FUNCTION_BLOCK "FB_BPSEthLink_V1.00"   // FB15, SCL
{ S7_Optimized_Access := 'TRUE' }
VERSION : 0.1
   VAR_INPUT
      IN_xBPSServerA : Bool;   // This istance is for BPS Server A
      IN_xCycleON : Bool;   // Cycle ON
      IN_xCycleONDel : Bool;   // Delayed cycle ON signal
      IN_xGeneralReset : Bool;   // General reset
      IN_xResetAlarms : Bool;   // Reset alarms
      IN_xFaultsEnabled : Bool;   // Faults enabled
      IN_xThisPLCActive : Bool;   // This PLC active
      IN_dLineSpeed_mm_min : DInt;   // Z301 speed [mm/min]
      IN_tStatusGeneral : Struct   // Status of general data
         dOptimizerMode : DInt;   // Optimizer mode (1=PLC 2=PC 3=Cullet)
         dExtOptSelected : DInt;   // External optimizer selected (1=PC A 2=PC B)
         dRibbonModality : DInt;   // Ribbon modality (1=Auto 4=Man)
         dAutoRibSelection : DInt;   // Automatic ribbon selection (0=Manual 1=Scanner 2=Camera)
         dTypeWanderSel : DInt;   // Wander type selection (1=Gross 2=Net)
         dActivePLC : DInt;   // Active PLC (1=PLC A 2=PLC B)
         dOptStatus : DInt;   // Status of optimizer connection (1=Disc 3=Conn 7=Anomaly)
         dScanStatus : DInt;   // Status of scanner connection (1=Disc 3=Conn 7=Anomaly)
         dScanGrossWidth_cmm : DInt;   // Scanner gross width [mm/100]
         dScanNetWidth_cmm : DInt;   // Scanner net width [mm/100]
         dScanGrossWander_cmm : DInt;   // Scanner gross wander [mm/100]
         dScanNetWander_cmm : DInt;   // Scanner net wander [mm/100]
         dCameraGrossWidth_cmm : DInt;   // Camera gross width [mm/100]
         dCameraNetWidth_cmm : DInt;   // Camera net width [mm/100]
         dCameraGrossWander_cmm : DInt;   // Camera gross wander [mm/100]
         dCameraNetWander_cmm : DInt;   // Camera net wander [mm/100]
         dWanderRecoveryThr_cmm : DInt;   // Wander recovery threshold [mm/100]
         dYC1WandRec_cmm : DInt;   // YCut 1 wander recovered [mm/100]
         dYC2WandRec_cmm : DInt;   // Ycut 2 wander recovered [mm/100]
      END_STRUCT;
      IN_tStatusEncoder : Struct   // Status of main tracking encoder
         dActualBTC_cmm : DInt;   // Actual BTC [mm/100]
         dTrackSpeed_mm_min : DInt;   // Tracking speed [mm/min]
         dActSelEnc : DInt;   // Actual selected encoder (1=Encoder#1 2=Encoder#2 4=Jog)
      END_STRUCT;
      IN_tStatusDigitizer_1 : Struct   // Status of digitizer_1
         dEncoderStatus : DInt;   // Encoder status (1=Stop 3=Running 7=Anomaly)
         dActualEncoderSpeed_mm_min : DInt;   // Actual encoder speed [mm/min]
         dDistanceSnapRoll_cmm : DInt;   // Distance from snaproll [mm/100]
      END_STRUCT;
      IN_tStatusDigitizer_2 : Struct   // Status of digitizer_2
         dEncoderStatus : DInt;   // Encoder status (1=Stop 3=Running 7=Anomaly)
         dActualEncoderSpeed_mm_min : DInt;   // Actual encoder speed [mm/min]
         dDistanceSnapRoll_cmm : DInt;   // Distance from snaproll [mm/100]
      END_STRUCT;
      IN_rgtStatusXCuts : Array[0.."DMAXXHEADS_IND"] of Struct   // Status of XCuts
         dDistanceFromSnaproll_cmm : DInt;   // Distance from snaproll [mm/100]
         dStatus : DInt;   // XCut actual status (1=Idle 3=Running 7=Faulted)
         dActualCarriagePos_cmm : DInt;   // XCut actual carriage position [mm/100]
         dXCutActualStatus : DInt;   // XCut actual status (1=Disabled 3=Enabled)
      END_STRUCT;
      IN_rgtStatusYCuts : Array[0.."DMAXYCUTBRIDGE_IND"] of Struct   // Status of YCut
         dDistanceSnapRoll_cmm : DInt;   // Distance from snaproll [mm/100]
         dBridgeStatus : DInt;   // Bridge actual status (1=OutOfProd 3=InProd 4=GlassBreak)
         rgxHeadProdOn : Array[0.."DMAXYHEADS_IND"] of Bool;   // Head#x production status
         rgxFireON : Array[0.."DMAXYHEADS_IND"] of Bool;   // Head#x fire status
         rgxArmON : Array[0.."DMAXYHEADS_IND"] of Bool;   // Head#x arm status
         rgdPosition_cmm : Array[0.."DMAXYHEADS_IND"] of DInt;   // Head#x position [mm/100]
      END_STRUCT;
      IN_rgtStatusMarkers : Array[0.."DMAXMARKERS_IND"] of Struct
         dDistanceFromSnaproll_cmm : DInt;   // Distance from snaproll [mm/100]
         dStatus : DInt;   // Marker actual status (1=Idle 3=Running 7=Faulted)
         dActualCarriagePos_cmm : DInt;   // Marker actual carriage position [mm/100]
         dMarkerActualStatus : DInt;   // Marker actual status (1=Disabled 3=Enabled)
      END_STRUCT;
      IN_tInterfaceID : Hw_Any;   // Interface ID BPS server A
      IN_tID : Conn_Ouc;   // Connection ID BPS server A
      IN_tRemoteAddress : IP_V4;   // Remote IP address BPS server A
      IN_uiRemotePort : UInt;   // Remote port BPS server A
   END_VAR
   VAR_IN_OUT
      INO_tCaps : "UDT_CapData_Tracking";   // Tracking plate DB
      INO_tInitialize : "GP_OB_Initialize";   // Service bits
      INO_tDefects : "UDT_DefectData_Tracking_Ext";   // Tracking defects
      INO_tMessages : "UDT_RP_TankMessages";   // Messages data
      INO_tAddMessageFromOpt : "UDT_RP_AddMessageCont_v2";   // Message add for received message
      INO_tRibbon : "UDT_RibbonData";   // Ribbon data
      INO_xMessageAnomaly : Bool;   // Message anomaly bit
   END_VAR
   VAR
      AUX_tCapToSend : "UDT_CapData";   // Cap data to send to BPS
      AUX_rgcPlateTelegram : Array[0..#DPLATETELEGRAMSIZE] of Char;   // Plate telegram container
      AUX_rgcStatusTelegram : Array[0..#DSTATUSTELEGRAMSIZE] of Char;   // Status telegram container
      AUX_rgcDefectTelegram : Array[0..#DDEFECTTELEGRAMSIZE] of Char;   // Defect telegram container
      AUX_rgcEventsTelegram : Array[0..#DEVENTSTELEGRAMSIZE] of Char;   // Events telegram container
      AUX_rgcRibbonTelegram : Array[0..#DRIBBONTELEGRAMSIZE] of Char;   // Ribbon telegram container
      AUX_dPlateTelegramNumByte : DInt;   // Number of byte on plate telegram
      AUX_dRibbonTelegramNumByte : DInt;   // Number of byte on ribbon telegram
      AUX_dStatusTelegramNumByte : DInt;   // Number of byte on status telegram
      AUX_dDefectTelegramNumByte : DInt;   // Number of byte on defect telegram
      AUX_dEventsTelegramNumByte : DInt;   // Number of byte on events telegram
      AUX_dLineSpeed_mm_min : DInt;   // Line speed z301
      ST_xRibbonTelegramAvail : Bool;   // Ribbon telegram available to send
      ST_xPlateTelegramAvail : Bool;   // Plate telegram available to send
      ST_xStatusTelegramAvail : Bool;   // Status telegram available to send
      ST_xDefectTelegramAvail : Bool;   // Defect telegram available to send
      ST_xEventsTelegramAvail : Bool;   // Events telegram available to send
      AUX_tStatusEncoder : Struct   // Status of main tracking encoder
         dActualBTC_cmm : DInt;   // Actual BTC [mm/100]
         dTrackSpeed_mm_min : DInt;   // Tracking speed [mm/min]
         dActSelEnc : DInt;   // Actual selected encoder (1=Encoder#1 2=Encoder#2 4=Jog)
      END_STRUCT;
      AUX_tStatusGeneral : Struct   // Status of general data
         dOptimizerMode : DInt;   // Optimizer mode (1=PLC 2=PC 3=Cullet)
         dExtOptSelected : DInt;   // External optimizer selected (1=PC A 2=PC B)
         dRibbonModality : DInt;   // Ribbon modality (1=Auto 4=Man)
         dAutoRibSelection : DInt;   // Automatic ribbon selection (0=Manual 1=Scanner 2=Camera)
         dTypeWanderSel : DInt;   // Wander type selection (1=Gross 2=Net)
         dActivePLC : DInt;   // Active PLC (1=PLC A 2=PLC B)
         dOptStatus : DInt;   // Status of optimizer connection (1=Disc 3=Conn 7=Anomaly)
         dScanStatus : DInt;   // Status of scanner connection (1=Disc 3=Conn 7=Anomaly)
         dScanGrossWidth_cmm : DInt;   // Scanner gross width [mm/100]
         dScanNetWidth_cmm : DInt;   // Scanner net width [mm/100]
         dScanGrossWander_cmm : DInt;   // Scanner gross wander [mm/100]
         dScanNetWander_cmm : DInt;   // Scanner net wander [mm/100]
         dCameraGrossWidth_cmm : DInt;   // Camera gross width [mm/100]
         dCameraNetWidth_cmm : DInt;   // Camera net width [mm/100]
         dCameraGrossWander_cmm : DInt;   // Camera gross wander [mm/100]
         dCameraNetWander_cmm : DInt;   // Camera net wander [mm/100]
         dWanderRecoveryThr_cmm : DInt;   // Wander recovery threshold [mm/100]
         dYC1WandRec_cmm : DInt;   // YCut 1 wander recovered [mm/100]
         dYC2WandRec_cmm : DInt;   // Ycut 2 wander recovered [mm/100]
      END_STRUCT;
      AUX_tStatusDigitizer_1 : Struct   // Status of digitizer_1
         dEncoderStatus : DInt;   // Encoder status (1=Stop 3=Running 7=Anomaly)
         dActualEncoderSpeed_mm_min : DInt;   // Actual encoder speed [mm/min]
         dDistanceSnapRoll_cmm : DInt;   // Distance from snaproll [mm/100]
      END_STRUCT;
      AUX_tStatusDigitizer_2 : Struct   // Status of digitizer_1
         dEncoderStatus : DInt;   // Encoder status (1=Stop 3=Running 7=Anomaly)
         dActualEncoderSpeed_mm_min : DInt;   // Actual encoder speed [mm/min]
         dDistanceSnapRoll_cmm : DInt;   // Distance from snaproll [mm/100]
      END_STRUCT;
      AUX_rgtStatusXCuts : Array[0.."DMAXXHEADS_IND"] of Struct   // Status of XCuts
         dDistanceFromSnaproll_cmm : DInt;   // Distance from snaproll [mm/100]
         dStatus : DInt;   // XCut actual status (1=Idle 3=Running 7=Faulted)
         dActualCarriagePos_cmm : DInt;   // XCut actual carriage position [mm/100]
         dXCutActualStatus : DInt;   // XCut actual status (1=Disabled 3=Enabled)
      END_STRUCT;
      AUX_rgtStatusMarkers : Array[0.."DMAXMARKERS_IND"] of Struct
         dDistanceFromSnaproll_cmm : DInt;   // Distance from snaproll [mm/100]
         dStatus : DInt;   // Marker actual status (1=Idle 3=Running 7=Faulted)
         dActualCarriagePos_cmm : DInt;   // Marker actual carriage position [mm/100]
         dMarkerActualStatus : DInt;   // Marker actual status (1=Disabled 3=Enabled)
      END_STRUCT;
      AUX_rgtStatusYCuts : Array[0.."DMAXYCUTBRIDGE_IND"] of Struct   // Status of YCut
         dDistanceSnapRoll_cmm : DInt;   // Distance from snaproll [mm/100]
         dBridgeStatus : DInt;   // Bridge actual status (1=OutOfProd 3=InProd 4=GlassBreak)
         rgxHeadProdOn : Array[0.."DMAXYHEADS_IND"] of Bool;   // Head#x production status
         rgxFireON : Array[0.."DMAXYHEADS_IND"] of Bool;   // Head#x fire status
         rgxArmON : Array[0.."DMAXYHEADS_IND"] of Bool;   // Head#x arm status
         rgdPosition_cmm : Array[0.."DMAXYHEADS_IND"] of DInt;   // Head#x position [mm/100]
      END_STRUCT;
      AUX_rgcSendTelegram : Array[0..#DSENDTELEGRAMSIZE] of Char;   // Send telegram buffer
      AUX_rgcRecvTelegram : Array[0..#DRECVTELEGRAMSIZE] of Char;   // Receive telegram
      AUX_rgcRecvBuffer : Array[0..#DRECVBUFFERSIZE] of Char;   // Receive buffer size
      AUX_dSendTelegramNumByte : DInt;   // Send telegram number of byte
      AUX_dNumByteRecvBuffer : DInt;   // Number of byte receive buffer
      AUX_rgcAnalyzedTelegram : Array[0..#DRECVTELEGRAMSIZE] of Char;   // Analyzed telegram
      AUX_rgcMetaData : Array[0..#DRECVTELEGRAMSIZE] of Char;   // Temp string with metadata
      tPhasesNetwork : Struct
         xSendBufferInProgress : Bool;   // Send data buffer in progress
         xEndSendBufferInProgress : Bool;   // End send data buffer in progress
         xSpare2 : Bool;
         xSpare3 : Bool;
         xSpare4 : Bool;
         xSpare5 : Bool;
         xSpare6 : Bool;
         xSpare7 : Bool;
         xSpare8 : Bool;
         xSpare9 : Bool;
         xSpare10 : Bool;
         xSpare11 : Bool;
         xSpare12 : Bool;
         xSpare13 : Bool;
         xSpare14 : Bool;
         xSpare15 : Bool;
         xSpare16 : Bool;
         xSpare17 : Bool;
         xSpare18 : Bool;
         xSpare19 : Bool;
         xSpare20 : Bool;
         xSpare21 : Bool;
         xSpare22 : Bool;
         xSpare23 : Bool;
         xSpare24 : Bool;
         xSpare25 : Bool;
         xSpare26 : Bool;
         xSpare27 : Bool;
         xSpare28 : Bool;
         xSpare29 : Bool;
         xSpare30 : Bool;
         xSpare31 : Bool;
      END_STRUCT;
      ST_xRetrySendTelegram : Bool;   // Retry send telegram
      ST_xPhasesInProgress : Bool;   // Phases in progress
      AUX_tConnData : TCON_IP_v4;   // Connection data structure
      AUX_xResetSendConnection : Bool;   // Reset send local connection
      FB_TSend : TSEND_C;   // Senda data
      FB_TRecv : TRCV_C;   // Receive data
      tALM : Struct   // HMI Alarms
         tS : Struct   // Stopping faults
            xTimeOutSendBPSData : Bool;   // Time out send BPS data
            xSpare_1 : Bool;
            xSpare_2 : Bool;
            xSpare_3 : Bool;
            xSpare_4 : Bool;
            xSpare_5 : Bool;
            xSpare_6 : Bool;
            xSpare_7 : Bool;
            xSpare_8 : Bool;
            xSpare_9 : Bool;
            xSpare_10 : Bool;
            xSpare_11 : Bool;
            xSpare_12 : Bool;
            xSpare_13 : Bool;
            xSpare_14 : Bool;
            xSpare_15 : Bool;
            xSpare_16 : Bool;
            xSpare_17 : Bool;
            xSpare_18 : Bool;
            xSpare_19 : Bool;
            xSpare_20 : Bool;
            xSpare_21 : Bool;
            xSpare_22 : Bool;
            xSpare_23 : Bool;
            xSpare_24 : Bool;
            xSpare_25 : Bool;
            xSpare_26 : Bool;
            xSpare_27 : Bool;
            xSpare_28 : Bool;
            xSpare_29 : Bool;
            xSpare_30 : Bool;
            xSpare_31 : Bool;
         END_STRUCT;
         tF : Struct   // Faults
            xSpare_0 : Bool;
            xSpare_1 : Bool;
            xSpare_2 : Bool;
            xSpare_3 : Bool;
            xSpare_4 : Bool;
            xSpare_5 : Bool;
            xSpare_6 : Bool;
            xSpare_7 : Bool;
            xSpare_8 : Bool;
            xSpare_9 : Bool;
            xSpare_10 : Bool;
            xSpare_11 : Bool;
            xSpare_12 : Bool;
            xSpare_13 : Bool;
            xSpare_14 : Bool;
            xSpare_15 : Bool;
            xSpare_16 : Bool;
            xSpare_17 : Bool;
            xSpare_18 : Bool;
            xSpare_19 : Bool;
            xSpare_20 : Bool;
            xSpare_21 : Bool;
            xSpare_22 : Bool;
            xSpare_23 : Bool;
            xSpare_24 : Bool;
            xSpare_25 : Bool;
            xSpare_26 : Bool;
            xSpare_27 : Bool;
            xSpare_28 : Bool;
            xSpare_29 : Bool;
            xSpare_30 : Bool;
            xSpare_31 : Bool;
         END_STRUCT;
         tW : Struct   // Warnings
            xSpare_0 : Bool;
            xSpare_1 : Bool;
            xSpare_2 : Bool;
            xSpare_3 : Bool;
            xSpare_4 : Bool;
            xSpare_5 : Bool;
            xSpare_6 : Bool;
            xSpare_7 : Bool;
            xSpare_8 : Bool;
            xSpare_9 : Bool;
            xSpare_10 : Bool;
            xSpare_11 : Bool;
            xSpare_12 : Bool;
            xSpare_13 : Bool;
            xSpare_14 : Bool;
            xSpare_15 : Bool;
            xSpare_16 : Bool;
            xSpare_17 : Bool;
            xSpare_18 : Bool;
            xSpare_19 : Bool;
            xSpare_20 : Bool;
            xSpare_21 : Bool;
            xSpare_22 : Bool;
            xSpare_23 : Bool;
            xSpare_24 : Bool;
            xSpare_25 : Bool;
            xSpare_26 : Bool;
            xSpare_27 : Bool;
            xSpare_28 : Bool;
            xSpare_29 : Bool;
            xSpare_30 : Bool;
            xSpare_31 : Bool;
         END_STRUCT;
      END_STRUCT;
      AUX_dPlateTelegramCounter : DInt := 1;   // Plate telegram counter
      AUX_dRibbonTelegramCounter : DInt := 1;   // Ribbon telegram counter
      AUX_dStatusTelegramCounter : DInt := 1;   // Status telegram counter
      AUX_dStatusServerCounter : DInt := 1;   // Status server counter
      AUX_dDefectTelegramCounter : DInt := 1;   // Defect telegram counter
      AUX_dEventsTelegramCounter : DInt := 1;   // Events telegram counter
      AUX_dWaitingNextStatus_ms : DInt;   // Waiting time for next status packet [ms]
      AUX_xResendAllPlate : Bool;   // Resend all plate after a disconnection
      AUX_xResendAllStatus : Bool;   // Resend all status after a disconnection
      AUX_tEmptyMessage : "UDT_RP_Message_v2";   // Empty message
      AUX_tRecvMessage : "UDT_RP_Message_v2";   // Received message
      AUX_rgstrMessageString : Array[0..#DMAXNUMSTR_IND] of String;
      AUX_rgstrSingleMexString : Array[0..#DMAXNUMSTR_IND] of String;
      AUX_tRibbonDataEl : "UDT_RibbonData_GlassData_SingleData";   // Ribbon data element
      AUX_rgxResendAllLastRib : Array[0.."DMAXGLASSDATAMACHINE_IND"] of Bool;   // Resend all last ribbon
   END_VAR
   VAR_TEMP
      TMP_dTail : DInt;
      TMP_xCapToSendFound : Bool;
      TMP_dIndex : DInt;
      TMP_uiNumChar : UInt;
      TMP_dLiteIndex : DInt;
      TMP_strTemp : String;
      TMP_dXCutIndex : DInt;
      TMP_dwValue : DWord;
      TMP_cValue : Char;
      TMP_strFixLite : String;
      TMP_dYCutIndex : DInt;
      TMP_strYCut : String;
      TMP_dYCutHeadIndex : DInt;
      TMP_strYCutIndex : String;
      TMP_strHeadIndex : String;
      TMP_strXCutIndex : String;
      TMP_strMarkerIndex : String;
      TMP_dIndexDef : DInt;
      TMP_strDefIndex : String;
      TMP_strDef : String;
      TMP_dCounter : DInt;
      TMP_dRemaining : DInt;
      TMP_iRetVal : Int;
      TMP_xSystemConnected : Bool;
      TMP_udCountString : UDInt;
      TMP_udPosition : UDInt;
      TMP_cSeparator : Char;
      TMP_cEndSeparator : Char;
      TMP_uiCount : UInt;
      TMP_dGlassDataIndex : DInt;
      TMP_xRibbonDataFound : Bool;
      TMP_dRibbonLastDataFound : DInt;
      TMP_dMarkerIndex : DInt;
      TMP_xThisBPSActive : Bool;
      TMP_dBridgeRequest : DInt;
      TMP_wBridgeMask : Word;
   END_VAR
   VAR CONSTANT
      BCONNTYPE : Byte := 16#0B;   // BPS Connection type
      DDELAYSTATUSPACKET_MS : DInt := 400;   // Status packet delay [ms]
      DMAXTELEGRAMCOUNTER : DInt := 2000000000;   // Maximum telegram counter
      DPLATETELEGRAMSIZE : DInt := 8192;   // Maximum plate telegram size
      DSTATUSTELEGRAMSIZE : DInt := 8192;   // Maximum status telegram size
      DDEFECTTELEGRAMSIZE : DInt := 8192;   // Maximum defect telegram size
      DEVENTSTELEGRAMSIZE : DInt := 8192;   // Maximum events telegram size
      DSENDTELEGRAMSIZE : DInt := 8192;   // Maximum size of the send telegram
      DRIBBONTELEGRAMSIZE : DInt := 1024;   // Maximum size of the ribbon telegram
      DRECVTELEGRAMSIZE : DInt := 1024;   // Maximum receive telegram size
      DRECVBUFFERSIZE : DInt := 8192;   // Maximum reveice buffer size
      DMAXMESSAGEPACKET : DInt := 20;   // Maximum number of message inside a packet
      STRSEPARATOR : Char := '|';   // Field separator
      STRPLATETELEGRAMID : Char := 'A';   // Plate telegram indentifier
      STR_CR : Char := '$R';   // CR
      STR_LF : Char := '$L';   // LF
      STRPLATETELCOUNTER : String := 'Z0=';
      STRCAPIDDESCR : String := 'Z1=';
      STRCAPHEADPOS : String := 'Z2=';
      STRCAPTAILPOS : String := 'Z3=';
      STRCAPLENGTH : String := 'Z4=';
      STRCAPWIDTH : String := 'Z5=';
      STRCAPTHICK : String := 'Z6=';
      STRCAPINDEX : String := 'Z7=';
      STRCAPFORMAT : String := 'Z8=';
      STRCAPNUMLITE : String := 'Z9=';
      STRCAPREQGAP : String := 'Z10=';
      STRCAPMAXCAP : String := 'Z11=';
      STRCAPCONVTOTLENGTH : String := 'Z12=';
      STRCAPGROSSWIDTH : String := 'Z13=';
      STRCAPNETWIDTH : String := 'Z14=';
      STRCAPIDEDGEOPSIDE : String := 'Z15=';
      STRCAPIDEDGEOPPOSIDE : String := 'Z16=';
      STRCAPWANDER : String := 'Z17=';
      STRCAPNETWANDER : String := 'Z18=';
      STRCAPGROSSWANDER : String := 'Z19=';
      STRCAPCOLOR : String := 'Z20=';
      STRCAPCOLORDESCR : String := 'Z21=';
      STRCAPSYSMEAS : String := 'Z22=';
      STRCAPYCUTBRIDGESEL : String := 'Z23=';
      STRCAPYCUTHEADNUM : String := 'Z24=';
      STRLITEIDENT : Char := 'A';
      STRLITEID : String := '1=';
      STRLITEPRODID : String := '2=';
      STRLITEPRODDESCR : String := '3=';
      STRLITEQUALID : String := '4=';
      STRLITEQUALDESCR : String := '5=';
      STRLITECAMERARECIPE : String := '6=';
      STRLITEWIDTH : String := '7=';
      STRLITEBARYCENTRE : String := '8=';
      STRLITECULLET : String := '9=';
      STRLITELAYERS : String := '10=';
      STRLITEMAINDEST : String := '11=';
      STRLITEALTDEST : String := '12=';
      STRLITE2NDDEST : String := '13=';
      STRLITESATPLATE : String := '14=';
      DPLATEARRAYLENGTH : DInt := 500;
      STRSTATUSTELEGRAMID : Char := 'B';
      STRSTATUSTELCOUNTER : String := 'TelegramCounter=';
      STRSTATUSSERVCOUNTER : String := 'ServerCounter=';
      STRSTATUSBTC : String := 'ActualEncoderValue=';
      STRSTATUSLEHRSPEED : String := 'ActualLehrSpeed=';
      STRSTATUSTRACKSPEED : String := 'ActualLineSpeed=';
      STRSTATUSACTSELENC : String := 'ActualSelEnc=';
      STRSTATUSDGT1STATUS : String := 'Digit1Status=';
      STRSTATUSDGT1SPEED : String := 'Digit1Speed=';
      STRSTATUSDGT1DISTSNAP : String := 'Digit1DistSnap=';
      STRSTATUSDGT2STATUS : String := 'Digit2Status=';
      STRSTATUSDGT2SPEED : String := 'Digit2Speed=';
      STRSTATUSDGT2DISTSNAP : String := 'Digit2DistSnap=';
      STRSTATUSXCUTDISTSNAP : String := 'DistSnapXCut';
      STRSTATUSXCUTSTATUS : String := 'StatusXCut';
      STRSTATUSXCUTACTPOS : String := 'ActPosXCut';
      STRSTATUSXCUTACTSTATUS : String := 'ActStatusXCut';
      STRSTATUSMARKDISTSNAP : String := 'DistSnapMark';
      STRSTATUSMARKSTATUS : String := 'StatusMark';
      STRSTATUSMARKACTPOS : String := 'ActPosXMark';
      STRSTATUSMARKACTSTATUS : String := 'ActStatusMark';
      STRSTATUSYCUT : String := 'YC';
      STRSTATUSYCUTPOS : String := '_HPos';
      STRSTATUSYCUTFIRE : String := '_HFire';
      STRSTATUSYCUTPROD : String := '_HProd';
      STRSTATUSYCUTARM : String := '_HArm';
      STRSTATUSYCUTSTATUS : String := '_BridgeStatus=';
      STRSTATUSYCUTSDISTSNAP : String := '_DistSnap=';
      STRSTATUSOPTSTATUS : String := 'OptimizerStatus=';
      STRSTATUSSCANNERSTATUS : String := 'ScannerStatus=';
      STRSTATUSACTIVEPLC : String := 'ActivePLC=';
      STRSTATUSRIBSELEC : String := 'AutomaticRibbonSelection=';
      STRSTATUSEXTOPTSEL : String := 'ExternalOptimizerSelected=';
      STRSTATUSOPTMODE : String := 'OptimizerMode=';
      STRSTATUSRIBMODE : String := 'RibbonModality=';
      STRSTATUSTYPEWANDER : String := 'TypeWanderSelection=';
      STRSTATUSSCANNERGROSSWIDTH : String := 'ScannerGrossWidth=';
      STRSTATUSSCANNERNETWIDTH : String := 'ScannerNetWidth=';
      STRSTATUSSCANNERGROSSWANDER : String := 'ScannerGrossWander=';
      STRSTATUSSCANNERNETWANDER : String := 'ScannerNetWander=';
      STRSTATUSCAMERAGROSSWIDTH : String := 'CameraGrossWidth=';
      STRSTATUSCAMERANETWIDTH : String := 'CameraNetWidth=';
      STRSTATUSCAMERAGROSSWANDER : String := 'CameraGrossWander=';
      STRSTATUSCAMERANETWANDER : String := 'CameraNetWander=';
      STRSTATUSWANDRECTHR : String := 'WanderRecoveryThreshold=';
      STRSTATUSWANDYC1 : String := 'YCut1_WanderRecovered=';
      STRSTATUSWANDYC2 : String := 'YCut2_WanderRecovered=';
      STRDEFECTTELEGRAMID : Char := 'C';
      STRDEFECTTELCOUNTER : String := 'Tc=';
      STRDEFECTNUMDEF : String := 'Nd=';
      STRDEFECTID : String := 'Id';
      STRDEFECTCLASS : String := 'Ca';
      STRDEFECTSUBTYPE : String := 'Sb';
      STRDEFECTXPOS : String := 'Xp';
      STRDEFECTYPOS : String := 'Yp';
      STRDEFECTTOTLENGTH : String := 'Tl';
      STRDEFECTTOTWIDTH : String := 'Tw';
      STRDEFECTCORELENGTH : String := 'Cl';
      STRDEFECTCOREWIDTH : String := 'Cw';
      STRDEFECTDISTLENGTH : String := 'Dl';
      STRDEFECTDISTWIDTH : String := 'Dw';
      STRDEFECTOPTVAL : String := 'Md';
      STRDEFECTSCID : String := 'Sd';
      STREVENTSTELEGRAMID : Char := 'D';
      STREVENTSTELCOUNTER : String := 'Tc=';
      STREVENTSCODE : String := 'Cd=';
      STREVENTSDATETIME : String := 'Dt=';
      STREVENTSIDENT : String := 'Id=';
      STREVENTSDATA1 : String := 'D1=';
      STREVENTSDATA2 : String := 'D2=';
      STREVENTSDATA3 : String := 'D3=';
      STREVENTSDATA4 : String := 'D4=';
      STREVENTSDATA5 : String := 'D5=';
      STREVENTSDATA6 : String := 'D6=';
      STREVENTSDATA7 : String := 'D7=';
      STREVENTSDATA8 : String := 'D8=';
      STREVENTSDATA9 : String := 'D9=';
      STREVENTSDATA10 : String := 'D10=';
      DMAXNUMSTR : DInt := 50;   // Maximum number of string on message
      DMAXNUMSTR_IND : DInt := 49;   // Maximum number of string on message index (Always -1)
      STRRIBBONTELEGRAMID : Char := 'F';   // Ribbon telegram ID
      STRRIBBONTELEGRAMCOUNT : String := 'Tc=';   // Ribbon telegram counter
      STRRIBBONSOURCEINDEX : String := 'Si=';   // Ribbon source index
      STRRIBBONLASTDATA : String := 'Ld=';   // Ribbon last data
      STRRIBBONGROSSWIDTH : String := 'Gw=';   // Ribbon gross width
      STRRIBBONNETWIDTH : String := 'Nw=';   // Ribbon net width
      STRRIBBONGROSSWANDER : String := 'Ga=';   // Ribbon gross wander
      STRRIBBONNETWANDER : String := 'Na=';   // Ribbon net wander
      STRRIBBONENCVALUE : String := 'En=';   // Ribbon encoder value
   END_VAR
BEGIN
   //---------- CHECK IF THERE ARE PLATE AVAILABLE FOR BPS -----------------------
   #TMP_xSystemConnected := TRUE;

   #TMP_xThisBPSActive := FALSE;

   IF #IN_xBPSServerA AND #IN_tStatusGeneral.dExtOptSelected = 1  THEN
        #TMP_xThisBPSActive := TRUE;
   ELSIF NOT #IN_xBPSServerA AND #IN_tStatusGeneral.dExtOptSelected = 2  THEN
       #TMP_xThisBPSActive := TRUE;
   END_IF;

   //If the connection is OFF resend all the information to BPS 
   IF #FB_TSend.s_TDIAG_Status.State <> b#16#04 THEN

       #AUX_xResendAllPlate := TRUE;
       #AUX_xResendAllStatus := TRUE;
       #ST_xRetrySendTelegram := FALSE;
       #ST_xPlateTelegramAvail := FALSE;
       #ST_xStatusTelegramAvail := FALSE;
       #ST_xEventsTelegramAvail := FALSE;

       IF (#IN_xBPSServerA AND #IN_tStatusGeneral.dExtOptSelected = 1) THEN
           #INO_tDefects.xBPSARequireAllDef := TRUE;
       END_IF;

       IF (NOT #IN_xBPSServerA AND #IN_tStatusGeneral.dExtOptSelected = 2) THEN
           #INO_tDefects.xBPSBRequireAllDef := TRUE;
       END_IF;

       #TMP_xSystemConnected := FALSE;

       FOR #TMP_dIndex := 0  TO "DMAXGLASSDATAMACHINE_IND" DO
           #AUX_rgxResendAllLastRib[#TMP_dIndex] := TRUE;
       END_FOR;


   END_IF;

   REGION BPS_RIBBON_TELEGRAM

   IF #TMP_xSystemConnected AND NOT #ST_xRibbonTelegramAvail THEN

       #TMP_xRibbonDataFound := FALSE;
       #TMP_dRibbonLastDataFound := 0;

       FOR #TMP_dGlassDataIndex := 0 TO #INO_tRibbon.dActualNumberGlassDataMachine - 1 DO

           //Check first the last data if has data
           IF (#INO_tRibbon.rgtGlassData[#TMP_dGlassDataIndex].tLastDataBuffer.xDataPresent AND 
               ((#INO_tRibbon.rgtGlassData[#TMP_dGlassDataIndex].tLastDataBuffer.xUpdateDataBPSA AND #IN_xBPSServerA) OR
                  (#AUX_rgxResendAllLastRib[#TMP_dGlassDataIndex]) OR         
                 (#INO_tRibbon.rgtGlassData[#TMP_dGlassDataIndex].tLastDataBuffer.xUpdateDataBPSB AND NOT #IN_xBPSServerA))) THEN

               #AUX_tRibbonDataEl := #INO_tRibbon.rgtGlassData[#TMP_dGlassDataIndex].tLastDataBuffer;

               #TMP_xRibbonDataFound := TRUE;
               #TMP_dRibbonLastDataFound := 1;

               IF #AUX_rgxResendAllLastRib[#TMP_dGlassDataIndex] = FALSE THEN

                   IF (#IN_xBPSServerA) THEN
                       #INO_tRibbon.rgtGlassData[#TMP_dGlassDataIndex].tLastDataBuffer.xUpdateDataBPSA := FALSE;
                   ELSE
                       #INO_tRibbon.rgtGlassData[#TMP_dGlassDataIndex].tLastDataBuffer.xUpdateDataBPSB := FALSE;
                   END_IF;

               END_IF;

               #AUX_rgxResendAllLastRib[#TMP_dGlassDataIndex] := FALSE;

               EXIT;

           END_IF;

           #TMP_dTail := #INO_tRibbon.rgtGlassData[#TMP_dGlassDataIndex].dBufferTail;

           //Search the element on the buffer
           WHILE (#TMP_dTail <> #INO_tRibbon.rgtGlassData[#TMP_dGlassDataIndex].dBufferHead) AND (#INO_tRibbon.rgtGlassData[#TMP_dGlassDataIndex].dBufferHead <> -1) DO

               //Increment the tail
               IF (#TMP_dTail + 1) >= "DMAXGLASSDATASECTORS" THEN
                   #TMP_dTail := 0;
               ELSE
                   #TMP_dTail+= 1;
               END_IF;

               IF (#INO_tRibbon.rgtGlassData[#TMP_dGlassDataIndex].rgtBuffer[#TMP_dTail].xDataPresent AND 
                   ((#INO_tRibbon.rgtGlassData[#TMP_dGlassDataIndex].rgtBuffer[#TMP_dTail].xUpdateDataBPSA AND #IN_xBPSServerA) OR        
                     (#INO_tRibbon.rgtGlassData[#TMP_dGlassDataIndex].rgtBuffer[#TMP_dTail].xUpdateDataBPSB AND NOT #IN_xBPSServerA))) THEN

                   #AUX_tRibbonDataEl := #INO_tRibbon.rgtGlassData[#TMP_dGlassDataIndex].rgtBuffer[#TMP_dTail];
                   #TMP_xRibbonDataFound := TRUE;

                   IF (#IN_xBPSServerA) THEN
                       #INO_tRibbon.rgtGlassData[#TMP_dGlassDataIndex].rgtBuffer[#TMP_dTail].xUpdateDataBPSA := FALSE;
                   ELSE
                       #INO_tRibbon.rgtGlassData[#TMP_dGlassDataIndex].rgtBuffer[#TMP_dTail].xUpdateDataBPSB := FALSE;
                   END_IF;

                   EXIT;
               END_IF;

           END_WHILE;

           IF #TMP_xRibbonDataFound THEN
               EXIT;
           END_IF;  

       END_FOR;

       //Prepare telegram for send the information to BPS            
       IF #TMP_xRibbonDataFound THEN

           #TMP_dIndex := 0;

           #AUX_rgcRibbonTelegram[#TMP_dIndex] := #STRRIBBONTELEGRAMID;
           #TMP_dIndex+=1;

           #AUX_rgcRibbonTelegram[#TMP_dIndex] := #STRSEPARATOR;
           #TMP_dIndex+=1;

           Strg_TO_Chars(Strg:= CONCAT_STRING(IN1 := #STRRIBBONTELEGRAMCOUNT ,IN2 := DINT_TO_STRING(#AUX_dRibbonTelegramCounter)),
               pChars:=#TMP_dIndex,
               Cnt=>#TMP_uiNumChar,
               Chars:=#AUX_rgcRibbonTelegram);
               #TMP_dIndex+=#TMP_uiNumChar;

           #AUX_rgcRibbonTelegram[#TMP_dIndex] := #STRSEPARATOR;
           #TMP_dIndex+=1;

           Strg_TO_Chars(Strg:= CONCAT_STRING(IN1 := #STRRIBBONSOURCEINDEX ,IN2 := DINT_TO_STRING(#TMP_dGlassDataIndex)),
               pChars:=#TMP_dIndex,
               Cnt=>#TMP_uiNumChar,
               Chars:=#AUX_rgcRibbonTelegram);
               #TMP_dIndex+=#TMP_uiNumChar;

           #AUX_rgcRibbonTelegram[#TMP_dIndex] := #STRSEPARATOR;
           #TMP_dIndex+=1;

           Strg_TO_Chars(Strg:= CONCAT_STRING(IN1 := #STRRIBBONLASTDATA ,IN2 := DINT_TO_STRING(#TMP_dRibbonLastDataFound)),
               pChars:=#TMP_dIndex,
               Cnt=>#TMP_uiNumChar,
               Chars:=#AUX_rgcRibbonTelegram);
               #TMP_dIndex+=#TMP_uiNumChar;

           #AUX_rgcRibbonTelegram[#TMP_dIndex] := #STRSEPARATOR;
           #TMP_dIndex+=1;

           Strg_TO_Chars(Strg:= CONCAT_STRING(IN1 := #STRRIBBONGROSSWIDTH ,IN2 := DINT_TO_STRING(#AUX_tRibbonDataEl.dGrossWidth_cmm)),
               pChars:=#TMP_dIndex,
               Cnt=>#TMP_uiNumChar,
               Chars:=#AUX_rgcRibbonTelegram);
               #TMP_dIndex+=#TMP_uiNumChar;

           #AUX_rgcRibbonTelegram[#TMP_dIndex] := #STRSEPARATOR;
           #TMP_dIndex+=1;

           Strg_TO_Chars(Strg:= CONCAT_STRING(IN1 := #STRRIBBONNETWIDTH ,IN2 := DINT_TO_STRING(#AUX_tRibbonDataEl.dNetWidth_cmm)),
               pChars:=#TMP_dIndex,
               Cnt=>#TMP_uiNumChar,
               Chars:=#AUX_rgcRibbonTelegram);
               #TMP_dIndex+=#TMP_uiNumChar;

           #AUX_rgcRibbonTelegram[#TMP_dIndex] := #STRSEPARATOR;
           #TMP_dIndex+=1;

           Strg_TO_Chars(Strg:= CONCAT_STRING(IN1 := #STRRIBBONGROSSWANDER ,IN2 := DINT_TO_STRING(#AUX_tRibbonDataEl.dGrossWander_cmm)),
               pChars:=#TMP_dIndex,
               Cnt=>#TMP_uiNumChar,
               Chars:=#AUX_rgcRibbonTelegram);
               #TMP_dIndex+=#TMP_uiNumChar;

           #AUX_rgcRibbonTelegram[#TMP_dIndex] := #STRSEPARATOR;
           #TMP_dIndex+=1;

           Strg_TO_Chars(Strg:= CONCAT_STRING(IN1 := #STRRIBBONNETWANDER ,IN2 := DINT_TO_STRING(#AUX_tRibbonDataEl.dNetWander_cmm)),
               pChars:=#TMP_dIndex,
               Cnt=>#TMP_uiNumChar,
               Chars:=#AUX_rgcRibbonTelegram);
               #TMP_dIndex+=#TMP_uiNumChar;

           #AUX_rgcRibbonTelegram[#TMP_dIndex] := #STRSEPARATOR;
           #TMP_dIndex+=1;

           Strg_TO_Chars(Strg:= CONCAT_STRING(IN1 := #STRRIBBONENCVALUE ,IN2 := DINT_TO_STRING(#AUX_tRibbonDataEl.dEncoderValue_cmm)),
               pChars:=#TMP_dIndex,
               Cnt=>#TMP_uiNumChar,
               Chars:=#AUX_rgcRibbonTelegram);
               #TMP_dIndex+=#TMP_uiNumChar;

           #AUX_rgcRibbonTelegram[#TMP_dIndex] := #STRSEPARATOR;
           #TMP_dIndex+=1;

           //Compile the number of byte and set telegram available to  send
           #AUX_rgcRibbonTelegram[#TMP_dIndex] := #STR_CR;
           #TMP_dIndex+=1;

           #AUX_rgcRibbonTelegram[#TMP_dIndex] := #STR_LF;

           #AUX_dRibbonTelegramNumByte := #TMP_dIndex + 1;

           IF #AUX_dRibbonTelegramCounter >= #DMAXTELEGRAMCOUNTER THEN
               #AUX_dRibbonTelegramCounter := 1;
           ELSE
               #AUX_dRibbonTelegramCounter += 1;
           END_IF;

           #ST_xRibbonTelegramAvail := TRUE;

       END_IF;

   END_IF;


   END_REGION 

   REGION BPS_EVENTS_TELEGRAM

   IF NOT #ST_xEventsTelegramAvail AND #TMP_xSystemConnected AND #TMP_xThisBPSActive (*AND FALSE*) THEN

       IF #INO_tMessages.dNumberOfMessage > 0  THEN

           #TMP_dCounter := 0;
           #TMP_dIndex := 0;

           WHILE (#TMP_dCounter < #DMAXMESSAGEPACKET) AND (#TMP_dCounter < #INO_tMessages.dNumberOfMessage) DO

               #AUX_rgcEventsTelegram[#TMP_dIndex] := #STREVENTSTELEGRAMID;
               #TMP_dIndex+=1;

               #AUX_rgcEventsTelegram[#TMP_dIndex] := #STRSEPARATOR;
               #TMP_dIndex+=1;

               Strg_TO_Chars(Strg:= CONCAT_STRING(IN1 := #STREVENTSTELCOUNTER ,IN2 := DINT_TO_STRING(#AUX_dEventsTelegramCounter)),
                             pChars:=#TMP_dIndex,
                             Cnt=>#TMP_uiNumChar,
                             Chars:=#AUX_rgcEventsTelegram);

               #TMP_dIndex+=#TMP_uiNumChar;

               #AUX_rgcEventsTelegram[#TMP_dIndex] := #STRSEPARATOR;
               #TMP_dIndex+=1;

               Strg_TO_Chars(Strg:= CONCAT_STRING(IN1 := #STREVENTSCODE ,IN2 := DINT_TO_STRING(#INO_tMessages.rgtMessages[#TMP_dCounter].dCodeEvent)),
                             pChars:=#TMP_dIndex,
                             Cnt=>#TMP_uiNumChar,
                             Chars:=#AUX_rgcEventsTelegram);

               #TMP_dIndex+=#TMP_uiNumChar;

               #AUX_rgcEventsTelegram[#TMP_dIndex] := #STRSEPARATOR;
               #TMP_dIndex+=1;





               Strg_TO_Chars(Strg:= CONCAT_STRING(IN1 := #STREVENTSDATETIME ,IN2 := "LGF_DTLtoString_ISO"("date":=#INO_tMessages.rgtMessages[#TMP_dCounter].dtDateTime, separator :='-')),
                             pChars:=#TMP_dIndex,
                             Cnt=>#TMP_uiNumChar,
                             Chars:=#AUX_rgcEventsTelegram);

               #TMP_dIndex+=#TMP_uiNumChar;

               #AUX_rgcEventsTelegram[#TMP_dIndex] := #STRSEPARATOR;
               #TMP_dIndex+=1;

               Strg_TO_Chars(Strg:= CONCAT_STRING(IN1 := #STREVENTSIDENT ,IN2 := #INO_tMessages.rgtMessages[#TMP_dCounter].strIdent),
                             pChars:=#TMP_dIndex,
                             Cnt=>#TMP_uiNumChar,
                             Chars:=#AUX_rgcEventsTelegram);

               #TMP_dIndex+=#TMP_uiNumChar;

               #AUX_rgcEventsTelegram[#TMP_dIndex] := #STRSEPARATOR;
               #TMP_dIndex+=1;

               Strg_TO_Chars(Strg:= CONCAT_STRING(IN1 := #STREVENTSDATA1 ,IN2 := DINT_TO_STRING(#INO_tMessages.rgtMessages[#TMP_dCounter].dEvent1)),
                             pChars:=#TMP_dIndex,
                             Cnt=>#TMP_uiNumChar,
                             Chars:=#AUX_rgcEventsTelegram);

               #TMP_dIndex+=#TMP_uiNumChar;

               #AUX_rgcEventsTelegram[#TMP_dIndex] := #STRSEPARATOR;
               #TMP_dIndex+=1;

               Strg_TO_Chars(Strg:= CONCAT_STRING(IN1 := #STREVENTSDATA2 ,IN2 := DINT_TO_STRING(#INO_tMessages.rgtMessages[#TMP_dCounter].dEvent2)),
                             pChars:=#TMP_dIndex,
                             Cnt=>#TMP_uiNumChar,
                             Chars:=#AUX_rgcEventsTelegram);

               #TMP_dIndex+=#TMP_uiNumChar;

               #AUX_rgcEventsTelegram[#TMP_dIndex] := #STRSEPARATOR;
               #TMP_dIndex+=1;

               Strg_TO_Chars(Strg:= CONCAT_STRING(IN1 := #STREVENTSDATA3 ,IN2 := DINT_TO_STRING(#INO_tMessages.rgtMessages[#TMP_dCounter].dEvent3)),
                             pChars:=#TMP_dIndex,
                             Cnt=>#TMP_uiNumChar,
                             Chars:=#AUX_rgcEventsTelegram);

               #TMP_dIndex+=#TMP_uiNumChar;

               #AUX_rgcEventsTelegram[#TMP_dIndex] := #STRSEPARATOR;
               #TMP_dIndex+=1;

               Strg_TO_Chars(Strg:= CONCAT_STRING(IN1 := #STREVENTSDATA4 ,IN2 := DINT_TO_STRING(#INO_tMessages.rgtMessages[#TMP_dCounter].dEvent4)),
                             pChars:=#TMP_dIndex,
                             Cnt=>#TMP_uiNumChar,
                             Chars:=#AUX_rgcEventsTelegram);

               #TMP_dIndex+=#TMP_uiNumChar;

               #AUX_rgcEventsTelegram[#TMP_dIndex] := #STRSEPARATOR;
               #TMP_dIndex+=1;

              Strg_TO_Chars(Strg:= CONCAT_STRING(IN1 := #STREVENTSDATA5 ,IN2 := DINT_TO_STRING(#INO_tMessages.rgtMessages[#TMP_dCounter].dEvent5)),
                             pChars:=#TMP_dIndex,
                             Cnt=>#TMP_uiNumChar,
                             Chars:=#AUX_rgcEventsTelegram);

               #TMP_dIndex+=#TMP_uiNumChar;

               #AUX_rgcEventsTelegram[#TMP_dIndex] := #STRSEPARATOR;
               #TMP_dIndex+=1;

              Strg_TO_Chars(Strg:= CONCAT_STRING(IN1 := #STREVENTSDATA6 ,IN2 := DINT_TO_STRING(#INO_tMessages.rgtMessages[#TMP_dCounter].dEvent6)),
                             pChars:=#TMP_dIndex,
                             Cnt=>#TMP_uiNumChar,
                             Chars:=#AUX_rgcEventsTelegram);

               #TMP_dIndex+=#TMP_uiNumChar;

               #AUX_rgcEventsTelegram[#TMP_dIndex] := #STRSEPARATOR;
               #TMP_dIndex+=1;

              Strg_TO_Chars(Strg:= CONCAT_STRING(IN1 := #STREVENTSDATA7 ,IN2 := DINT_TO_STRING(#INO_tMessages.rgtMessages[#TMP_dCounter].dEvent7)),
                             pChars:=#TMP_dIndex,
                             Cnt=>#TMP_uiNumChar,
                             Chars:=#AUX_rgcEventsTelegram);

               #TMP_dIndex+=#TMP_uiNumChar;

               #AUX_rgcEventsTelegram[#TMP_dIndex] := #STRSEPARATOR;
               #TMP_dIndex+=1;

              Strg_TO_Chars(Strg:= CONCAT_STRING(IN1 := #STREVENTSDATA8 ,IN2 := DINT_TO_STRING(#INO_tMessages.rgtMessages[#TMP_dCounter].dEvent8)),
                             pChars:=#TMP_dIndex,
                             Cnt=>#TMP_uiNumChar,
                             Chars:=#AUX_rgcEventsTelegram);

               #TMP_dIndex+=#TMP_uiNumChar;

               #AUX_rgcEventsTelegram[#TMP_dIndex] := #STRSEPARATOR;
               #TMP_dIndex+=1;

              Strg_TO_Chars(Strg:= CONCAT_STRING(IN1 := #STREVENTSDATA9 ,IN2 := DINT_TO_STRING(#INO_tMessages.rgtMessages[#TMP_dCounter].dEvent9)),
                             pChars:=#TMP_dIndex,
                             Cnt=>#TMP_uiNumChar,
                             Chars:=#AUX_rgcEventsTelegram);

               #TMP_dIndex+=#TMP_uiNumChar;

               #AUX_rgcEventsTelegram[#TMP_dIndex] := #STRSEPARATOR;
               #TMP_dIndex+=1;

              Strg_TO_Chars(Strg:= CONCAT_STRING(IN1 := #STREVENTSDATA10 ,IN2 := DINT_TO_STRING(#INO_tMessages.rgtMessages[#TMP_dCounter].dEvent10)),
                             pChars:=#TMP_dIndex,
                             Cnt=>#TMP_uiNumChar,
                             Chars:=#AUX_rgcEventsTelegram);

               #TMP_dIndex+=#TMP_uiNumChar;

               #AUX_rgcEventsTelegram[#TMP_dIndex] := #STRSEPARATOR;
               #TMP_dIndex+=1;

               //Compile the number of byte and set telegram available to  send
               #AUX_rgcEventsTelegram[#TMP_dIndex] := #STR_CR;
               #TMP_dIndex+=1;

               #AUX_rgcEventsTelegram[#TMP_dIndex] := #STR_LF;
               #TMP_dIndex+=1;

               IF #AUX_dEventsTelegramCounter >= #DMAXTELEGRAMCOUNTER THEN
                   #AUX_dEventsTelegramCounter := 1;
               ELSE
                   #AUX_dEventsTelegramCounter += 1;
               END_IF;

               #INO_tMessages.rgtMessages[#TMP_dCounter] := #AUX_tEmptyMessage;

               #TMP_dCounter+= 1;

           END_WHILE;

           #AUX_dEventsTelegramNumByte := #TMP_dIndex;
           #ST_xEventsTelegramAvail := TRUE;

           #TMP_dRemaining := #INO_tMessages.dNumberOfMessage - #TMP_dCounter;

           IF #TMP_dRemaining > 0 THEN
               #TMP_iRetVal :=  MOVE_BLK_VARIANT(   SRC:=#INO_tMessages.rgtMessages, 
                                   COUNT:=DINT_TO_UDINT(#TMP_dRemaining), 
                                   SRC_INDEX:=#TMP_dCounter, 
                                   DEST_INDEX:=0, 
                                   DEST=>#INO_tMessages.rgtMessages);
               //Reset the remaining
               FOR #TMP_dIndex := #TMP_dRemaining TO #INO_tMessages.dNumberOfMessage - 1 DO
                   #INO_tMessages.rgtMessages[#TMP_dIndex] := #AUX_tEmptyMessage;
               END_FOR;

               #INO_tMessages.dNumberOfMessage := #TMP_dRemaining;

           ELSE
               #INO_tMessages.dNumberOfMessage := 0;
           END_IF;
       END_IF;
   END_IF;

   END_REGION BPS_EVENTS_TELEGRAM

   REGION BPS_DEFECTS_TELEGRAM

   IF NOT #ST_xDefectTelegramAvail AND #TMP_xSystemConnected AND #TMP_xThisBPSActive THEN

       IF #INO_tDefects.tDefectsForReport.dNumberOfDefect > 0 THEN

           #TMP_dIndex := 0;

           #AUX_rgcDefectTelegram[#TMP_dIndex] := #STRDEFECTTELEGRAMID;
           #TMP_dIndex+=1;

           #AUX_rgcDefectTelegram[#TMP_dIndex] := #STRSEPARATOR;
           #TMP_dIndex+=1;

           Strg_TO_Chars(Strg:= CONCAT_STRING(IN1 := #STRDEFECTTELCOUNTER ,IN2 := DINT_TO_STRING(#AUX_dDefectTelegramCounter)),
                         pChars:=#TMP_dIndex,
                         Cnt=>#TMP_uiNumChar,
                         Chars:=#AUX_rgcDefectTelegram);

           #TMP_dIndex+=#TMP_uiNumChar;

           #AUX_rgcDefectTelegram[#TMP_dIndex] := #STRSEPARATOR;
           #TMP_dIndex+=1;

           Strg_TO_Chars(Strg:= CONCAT_STRING(IN1 := #STRDEFECTNUMDEF ,IN2 := DINT_TO_STRING(#INO_tDefects.tDefectsForReport.dNumberOfDefect)),
                         pChars:=#TMP_dIndex,
                         Cnt=>#TMP_uiNumChar,
                         Chars:=#AUX_rgcDefectTelegram);

           #TMP_dIndex+=#TMP_uiNumChar;

           #AUX_rgcDefectTelegram[#TMP_dIndex] := #STRSEPARATOR;
           #TMP_dIndex+=1;

           FOR #TMP_dIndexDef := 0 TO #INO_tDefects.tDefectsForReport.dNumberOfDefect - 1 DO

               #TMP_strDefIndex := DINT_TO_STRING(#TMP_dIndexDef + 1);   

               #TMP_strDefIndex := DELETE(IN:=#TMP_strDefIndex, L:=1, P:=1);

               //Defect ID
               #TMP_strDef := CONCAT_STRING(IN1 := #STRDEFECTID ,IN2 := #TMP_strDefIndex);
               #TMP_strDef := CONCAT_STRING(IN1 := #TMP_strDef,IN2 := '=');

               Strg_TO_Chars(Strg:= CONCAT_STRING(IN1 := #TMP_strDef ,IN2 := DINT_TO_STRING(#INO_tDefects.tDefectsForReport.rgtDefects[#TMP_dIndexDef].dID)),
                         pChars:=#TMP_dIndex,
                         Cnt=>#TMP_uiNumChar,
                         Chars:=#AUX_rgcDefectTelegram);
               #TMP_dIndex+=#TMP_uiNumChar;

               #AUX_rgcDefectTelegram[#TMP_dIndex] := #STRSEPARATOR;
               #TMP_dIndex+=1;

               //Defect class
               #TMP_strDef := CONCAT_STRING(IN1 := #STRDEFECTCLASS ,IN2 := #TMP_strDefIndex);
               #TMP_strDef := CONCAT_STRING(IN1 := #TMP_strDef,IN2 := '=');

               Strg_TO_Chars(Strg:= CONCAT_STRING(IN1 := #TMP_strDef ,IN2 := DINT_TO_STRING(#INO_tDefects.tDefectsForReport.rgtDefects[#TMP_dIndexDef].dClass)),
                         pChars:=#TMP_dIndex,
                         Cnt=>#TMP_uiNumChar,
                         Chars:=#AUX_rgcDefectTelegram);
               #TMP_dIndex+=#TMP_uiNumChar;

               #AUX_rgcDefectTelegram[#TMP_dIndex] := #STRSEPARATOR;
               #TMP_dIndex+=1;

               //Defect subtype
               #TMP_strDef := CONCAT_STRING(IN1 := #STRDEFECTSUBTYPE ,IN2 := #TMP_strDefIndex);
               #TMP_strDef := CONCAT_STRING(IN1 := #TMP_strDef,IN2 := '=');

               Strg_TO_Chars(Strg:= CONCAT_STRING(IN1 := #TMP_strDef ,IN2 := DINT_TO_STRING(#INO_tDefects.tDefectsForReport.rgtDefects[#TMP_dIndexDef].dSubType)),
                         pChars:=#TMP_dIndex,
                         Cnt=>#TMP_uiNumChar,
                         Chars:=#AUX_rgcDefectTelegram);
               #TMP_dIndex+=#TMP_uiNumChar;

               #AUX_rgcDefectTelegram[#TMP_dIndex] := #STRSEPARATOR;
               #TMP_dIndex+=1;

               //Defect XPOS
               #TMP_strDef := CONCAT_STRING(IN1 := #STRDEFECTXPOS ,IN2 := #TMP_strDefIndex);
               #TMP_strDef := CONCAT_STRING(IN1 := #TMP_strDef,IN2 := '=');

               Strg_TO_Chars(Strg:= CONCAT_STRING(IN1 := #TMP_strDef ,IN2 := DINT_TO_STRING(#INO_tDefects.tDefectsForReport.rgtDefects[#TMP_dIndexDef].dXPosition_cmm)),
                         pChars:=#TMP_dIndex,
                         Cnt=>#TMP_uiNumChar,
                         Chars:=#AUX_rgcDefectTelegram);
               #TMP_dIndex+=#TMP_uiNumChar;

               #AUX_rgcDefectTelegram[#TMP_dIndex] := #STRSEPARATOR;
               #TMP_dIndex+=1;

               //Defect YPOS
               #TMP_strDef := CONCAT_STRING(IN1 := #STRDEFECTYPOS ,IN2 := #TMP_strDefIndex);
               #TMP_strDef := CONCAT_STRING(IN1 := #TMP_strDef,IN2 := '=');

               Strg_TO_Chars(Strg:= CONCAT_STRING(IN1 := #TMP_strDef ,IN2 := DINT_TO_STRING(#INO_tDefects.tDefectsForReport.rgtDefects[#TMP_dIndexDef].dYPosition_cmm)),
                         pChars:=#TMP_dIndex,
                         Cnt=>#TMP_uiNumChar,
                         Chars:=#AUX_rgcDefectTelegram);
               #TMP_dIndex+=#TMP_uiNumChar;

               #AUX_rgcDefectTelegram[#TMP_dIndex] := #STRSEPARATOR;
               #TMP_dIndex+=1;

               //Defect Tot length
               #TMP_strDef := CONCAT_STRING(IN1 := #STRDEFECTTOTLENGTH ,IN2 := #TMP_strDefIndex);
               #TMP_strDef := CONCAT_STRING(IN1 := #TMP_strDef,IN2 := '=');

               Strg_TO_Chars(Strg:= CONCAT_STRING(IN1 := #TMP_strDef ,IN2 := DINT_TO_STRING(#INO_tDefects.tDefectsForReport.rgtDefects[#TMP_dIndexDef].dTotalLength_um)),
                         pChars:=#TMP_dIndex,
                         Cnt=>#TMP_uiNumChar,
                         Chars:=#AUX_rgcDefectTelegram);
               #TMP_dIndex+=#TMP_uiNumChar;

               #AUX_rgcDefectTelegram[#TMP_dIndex] := #STRSEPARATOR;
               #TMP_dIndex+=1;

               //Defect Tot width
               #TMP_strDef := CONCAT_STRING(IN1 := #STRDEFECTTOTWIDTH ,IN2 := #TMP_strDefIndex);
               #TMP_strDef := CONCAT_STRING(IN1 := #TMP_strDef,IN2 := '=');

               Strg_TO_Chars(Strg:= CONCAT_STRING(IN1 := #TMP_strDef ,IN2 := DINT_TO_STRING(#INO_tDefects.tDefectsForReport.rgtDefects[#TMP_dIndexDef].dTotalWidth_um)),
                         pChars:=#TMP_dIndex,
                         Cnt=>#TMP_uiNumChar,
                         Chars:=#AUX_rgcDefectTelegram);
               #TMP_dIndex+=#TMP_uiNumChar;

               #AUX_rgcDefectTelegram[#TMP_dIndex] := #STRSEPARATOR;
               #TMP_dIndex+=1;

               //Defect Tot width
               #TMP_strDef := CONCAT_STRING(IN1 := #STRDEFECTTOTWIDTH ,IN2 := #TMP_strDefIndex);
               #TMP_strDef := CONCAT_STRING(IN1 := #TMP_strDef,IN2 := '=');

               Strg_TO_Chars(Strg:= CONCAT_STRING(IN1 := #TMP_strDef ,IN2 := DINT_TO_STRING(#INO_tDefects.tDefectsForReport.rgtDefects[#TMP_dIndexDef].dTotalWidth_um)),
                         pChars:=#TMP_dIndex,
                         Cnt=>#TMP_uiNumChar,
                         Chars:=#AUX_rgcDefectTelegram);
               #TMP_dIndex+=#TMP_uiNumChar;

               #AUX_rgcDefectTelegram[#TMP_dIndex] := #STRSEPARATOR;
               #TMP_dIndex+=1;

               //Defect core length
               #TMP_strDef := CONCAT_STRING(IN1 := #STRDEFECTCORELENGTH ,IN2 := #TMP_strDefIndex);
               #TMP_strDef := CONCAT_STRING(IN1 := #TMP_strDef,IN2 := '=');

               Strg_TO_Chars(Strg:= CONCAT_STRING(IN1 := #TMP_strDef ,IN2 := DINT_TO_STRING(#INO_tDefects.tDefectsForReport.rgtDefects[#TMP_dIndexDef].dCoreLength_um)),
                         pChars:=#TMP_dIndex,
                         Cnt=>#TMP_uiNumChar,
                         Chars:=#AUX_rgcDefectTelegram);
               #TMP_dIndex+=#TMP_uiNumChar;

               #AUX_rgcDefectTelegram[#TMP_dIndex] := #STRSEPARATOR;
               #TMP_dIndex+=1;

               //Defect core width
               #TMP_strDef := CONCAT_STRING(IN1 := #STRDEFECTCOREWIDTH ,IN2 := #TMP_strDefIndex);
               #TMP_strDef := CONCAT_STRING(IN1 := #TMP_strDef,IN2 := '=');